VERSION : 1.2
// ellipse_C calculates the circumference of an ellipe based on the two radians R1 and R2
   VAR_INPUT
      R1 : Real;
      R2 : Real;
   END_VAR
BEGIN


   #ELLIPSE_C := "PI" * (3.0 * (#R1+#R2) - SQRT((3.0 * #R1 + #R2) * (3.0 * #R2 + #R1)));


   (* revision histroy
   hm  16. oct 2007    rev 1.0
       original version

   hm  18. oct. 2008   rev 1.1
       using math constants

   hm  10. mar. 2009   rev 1.2
       changed syntax of real constants to 0.0

   *)
END_FUNCTION

FUNCTION "SPHERE_V" : Real   // FC160, SCL
TITLE = SPHERE_V
{ S7_Optimized_Access := 'FALSE' }
AUTHOR : hugo
FAMILY : GEOMETRY
NAME : SPHERE_V
VERSION : 1.2
// sphere_V calculates the Volume of a Sphere
   VAR_INPUT
      rx : Real;
   END_VAR
BEGIN


     #SPHERE_V := 4.188790205 * #rx * #rx * #rx;

   (* revision histroy
   hm  16. oct 2007  rev 1.0
     original version

   hm  4. dec 2007   rev 1.1
     changed code for better performance

   hm  22. feb 2008    rev 1.2
     changed code for better performance
   *)
END_FUNCTION

FUNCTION "TRIANGLE_A" : Real   // FC161, SCL
TITLE = TRIANGLE_A
{ S7_Optimized_Access := 'FALSE' }
AUTHOR : hugo
FAMILY : GEOMETRY
NAME : TRIANG_A
VERSION : 1.2
// triangle_A calculates the Area of a triangle.
// if any input is 0 it will be neglected and the are will be calculated from eiter:
// two sides and an angle (s1 and S2 and the angle A1) or 3 sides.
// 
// uses: RAD [FC100]
//       MODR [FC97] 
//       FLOOR2 [FC82]
   VAR_INPUT
      S1 : Real;
      "A" : Real;
      S2 : Real;
      S3 : Real;
   END_VAR
BEGIN


   IF #"A" = 0.0 THEN
       #TRIANGLE_A := SQRT((#S1+#S2+#S3) * (#S1+#S2-#S3) * (#S2+#S3-#S1) * (#S3+#S1-#S2)) * 0.25;
   ELSE
       #TRIANGLE_A := #S1 * #S2 * SIN("RAD"(#"A")) * 0.5;
   END_IF;


   (* revision histroy
   hm  16. oct 2007    rev 1.0
       original version

   hm  22. feb 2008    rev 1.1
       improved performance

   hm  10. mar. 2009   rev 1.2
       changed syntax of real constants to 0.0

   *)
END_FUNCTION

FUNCTION "CIRCLE_SEG" : Real   // FC428, SCL
TITLE = CIRCLE_SEG
{ S7_Optimized_Access := 'FALSE' }
AUTHOR : hugo
FAMILY : GEOMETRY
NAME : CIRCLSEG
VERSION : 1.0
// CIRCLE_SEG calculates the Area of a circle segement enclosed between a sectant line and the circumference.
   VAR_INPUT
      RX : Real;
      HX : Real;
   END_VAR
BEGIN


   IF #RX > 0.0 THEN
     #CIRCLE_SEG := 2.0 * ACOS(1.0 - LIMIT(MN:=0.0,IN:=#HX / #RX,MX:=2.0));
     #CIRCLE_SEG := (#CIRCLE_SEG - SIN(#CIRCLE_SEG)) *#RX * #RX / 2.0;
   END_IF;


   (* revision histroy
   hm  10. mar 2010  rev 1.0
     original version

   *)
END_FUNCTION

// ===== PLC "Mathematical functions"  Unspecific CPU S7 300 =====

VAR_GLOBAL CONSTANT   // PLC tag table "STEP7 classic symbols"
   "debug" : Bool := FALSE;
   "N" : Int := 0;
   "offset" : Int := 0;
   "offset_1" : DWord := 0;
END_VAR

TYPE "XY_LINEAR_INT"
VERSION : 0.0
   STRUCT
      XY : Array[1..20, 0..1] of Real;
   END_STRUCT;
END_TYPE

TYPE "XY_POLYNOM_INT"
VERSION : 0.0
   STRUCT
      XY : Array[1..5, 0..1] of Real;
   END_STRUCT;
END_TYPE

TYPE "C_F_POLY"
VERSION : 0.0
   STRUCT
      C : Array[0..7] of Real;
   END_STRUCT;
END_TYPE

DATA_BLOCK "IDB_STIME"   // DB64
{ S7_Optimized_Access := 'FALSE' }
AUTHOR : dalbi
FAMILY : MEASURE
VERSION : 0.0
// stored: InstanceOfName STIME
"STIME"
BEGIN
END_DATA_BLOCK

FUNCTION_BLOCK "FT_AVG"   // FB23, SCL
TITLE = FT_AVG
{ S7_Optimized_Access := 'FALSE' }
AUTHOR : hugo
FAMILY : FUNCT
NAME : FT_AVG
VERSION : 1.5
// this function calculates the average over n samples from a sequential input
// the input values are shifted into an N deep buffer and the avg of this buffer is diplayed at anytime on the output.
// a rst will load the buffer with the current in value..
//  
// uses: DELAY [FB107]
//       INC1 [FC53]
   VAR_INPUT
      IN : Real;
      "E" : Bool := TRUE;
      N : Int := 32;
      RST : Bool;
   END_VAR
   VAR_OUTPUT
      AVG : Real;
   END_VAR
   VAR
      buff : "DELAY";
      i : Int;
      init : Bool;
   END_VAR
BEGIN


   (* limit n to a max of 32 because delay can do max 32 cycles *)
   #buff.N := LIMIT(MN:=0,IN:=#N,MX:=32);

   IF NOT #init OR #RST THEN
       FOR #i := 1 TO #N DO
           #buff(IN := #IN);
       END_FOR;
       #AVG := #IN;
       #init := TRUE;
   ELSIF #"E" THEN
       #buff(IN := #IN);
       #AVG := #AVG + (#IN - #buff.OUT) / INT_TO_REAL(#N);
   END_IF;


   (* revision history

   hm  7. jan. 2007    rev 1.1
       chaged rst logic to load the buffer with the actual input value instead of 0.
       added en input to allow better control of signal flow
       added init to load the buffer with in at startup to avoid rampup at beginning.
       deleted unused variable cnt.

   hm  14. jun. 2008   rev 1.2
       set default for input en = TRUE and N = 32

   hm  10. oct. 2008   rev 1.3
       improved performance

   hm  18. oct. 2008   rev 1.4
       changed input en to e for compatibility reasons

   hm  10. mar. 2009   rev 1.5
       added type conversion for compatibility reasons

   *)
END_FUNCTION_BLOCK

FUNCTION_BLOCK "FT_MIN_MAX"   // FB24, SCL
TITLE = FT_MIN_MAX
{ S7_Optimized_Access := 'FALSE' }
AUTHOR : hugo
FAMILY : FUNCT
NAME : MIN_MAX
VERSION : 1.0
// this function block stores the min and max value of an input signal.
// when rst is true the mn and mx outputs are set to the in value.
// when a rst is never active the function autoresets to the in value at startup.
// since the input might not be present at first cycle the mn and mx are set during second cycle.
   VAR_INPUT
      in : Real;
      rst : Bool;
   END_VAR
   VAR_OUTPUT
      mx : Real;
      mn : Real;
   END_VAR
   VAR
      init : Bool;
   END_VAR
BEGIN


     IF #rst OR NOT #init THEN
       #mn := #in;
       #mx := #in;
       #init := 1;
     ELSIF #in < #mn THEN
       #mn := #in;
     ELSIF #in > #mx THEN 
       #mx := #in;
     END_IF;
END_FUNCTION_BLOCK

FUNCTION_BLOCK "FT_RMP"   // FB25, SCL
TITLE = FT_RMP
{ S7_Optimized_Access := 'FALSE' }
AUTHOR : oscat
FAMILY : FUNCT
NAME : RMP
VERSION : 1.4
// this ramp function follows an input signal with a linear ramp up or down, the up or down speed can be set with KF and KR.
// a K factor of 1 means 1 unit per second on the output. K factors can only be positive and not negative.
// a busy output signals the ramp is running or busy false means the in value is present on the output.
// a rmp input false means the output follows the input dierctly while a rmp = true means the output follows the input with a ramp.
// a updn output signal the directon of the ramp (up or down).
// 
// uses: T_PLC_MS [FC64]
//       STIME [FB64],IDB_STIME [DB64]
   VAR_INPUT
      Rmp : Bool := TRUE;
      in : Real;
      KR : Real;
      KF : Real;
   END_VAR
   VAR_OUTPUT
      out : Real;
      busy : Bool;
      UD : Bool;
   END_VAR
   VAR
      tx : Time;
      last : Time;
      init : Bool;
   END_VAR
BEGIN


     (* read system time *)
     #tx := T_CONV(DWORD_TO_DINT("T_PLC_MS"())) - #last;

     IF NOT #init THEN
       #init := TRUE;
       #last := #tx;
       #tx := t#0s;
       #out := #in;
     END_IF;
     IF NOT #Rmp THEN
       #out := #in;
       #busy := FALSE;
     ELSIF #out > #in THEN
       (* ramp down *)
       #out := #out - DINT_TO_REAL(T_CONV(#tx)) * 0.001 * #KF;
       #out := MAX(IN1:=#in,IN2:=#out);
     ELSIF #out < #in THEN
       (* ramp up *)
       #out := #out + DINT_TO_REAL(T_CONV(#tx)) * 0.001 * #KR;
       #out := MIN(IN1:=#in,IN2:=#out);
     END_IF;

     (* set busy and dir flags *)
     IF #out < #in THEN
       #busy := TRUE;
       #UD := 1;
     ELSIF #out > #in THEN
       #busy := TRUE;
       #UD := 0;
     ELSE
       #busy := FALSE;
     END_IF;
     #last := #last + #tx;


   (* revision history:

   hm 8.10.2006      rev 1.1
     added ud output

   hm 12. feb 2007   rev 1.2
     added init variable and corrected a possible startup problem

   hm  17. sep 2007  rev 1.3
     replaced time() with t_plc_ms() for compatibility reasons

   hm  25. jan 2008  rev 1.4
     performance improvements
     allow KR and KF to be 0
   *)
END_FUNCTION_BLOCK

FUNCTION_BLOCK "STIME"   // FB64, SCL
TITLE = STIME
{ S7_Optimized_Access := 'FALSE' }
AUTHOR : dalbi
FAMILY : MEASURE
NAME : STIME
VERSION : 1.4
// this function block makes sure that the timer of a siemens sps counts from 0 - 2^32-1.
   VAR_OUTPUT
      tx : DWord;
      at_tx AT tx : Array[0..31] of Bool;
   END_VAR
   VAR
      last_time : DWord;
      bit31 : Bool;
      init : Bool := TRUE;
   END_VAR
   VAR_TEMP
      TOP_SI : Struct
         EV_CLASS : Byte;
         EV_NUM : Byte;
         PRIORITY : Byte;
         NUM : Byte;
         TYP2_3 : Byte;
         TYP1 : Byte;
         ZI1 : Word;
         ZI2_3 : DWord;
      END_STRUCT;
      START_UP_SI : Struct
         EV_CLASS : Byte;
         EV_NUM : Byte;
         PRIORITY : Byte;
         NUM : Byte;
         TYP2_3 : Byte;
         TYP1 : Byte;
         ZI1 : Word;
         ZI2_3 : DWord;
      END_STRUCT;
      ERR : Int;
   END_VAR
BEGIN


   (* this FB is only necessary for siemens sps
   the siemens sps timer counts from 0 to 2^31-1 and starts at 0 sfter overrun.
   this means that the bit 31 (the highest bit ) will never be used and therefore
   a problem arises when t2 - t1 is checked.
   t2 - t1 is always valid also in an timer overrun situation where the time t1 is very high and t2 is very low.
   the result of the subtraction t2 - t1 however is still valid.
   this calculation does not work for soiemens because the highest bit is not used.

   this module stores the highest bit, changes the highest bit at every overrun occurence and stuffs ther highest bit in the output.
   the output is then used by t_plc_us and t_plc_ms.

   the correction needs and fb and not a function because the value of the highest bit has to be stored.

   do never use this function block in a codesys environment. the timer in codesys is correct and runs from 0 to 2^32-1
   *)

   (* read actual startup info *)
   (* OB1_SCAN_1  BYTE  -  B#16#01: Abschluss des Neustarts (Warmstarts)
                        -  B#16#02: Abschluss des Wiederanlaufs
                        -  B#16#03: Abschluss des freien Zyklus
                        -  B#16#04: Abschluss des Kaltstarts
                        -  B#16#05: Erster OB 1-Zyklus der neuen Master-CPU nach 
                                    Master-Reserve-Umschaltung und STOP des 
                                    bisherigen Masters *)

   #ERR := RD_SINFO (TOP_SI => #TOP_SI, START_UP_SI => #START_UP_SI);

   (* reset last_time on system startup *)
   IF #TOP_SI.EV_NUM = 1 OR #TOP_SI.EV_NUM = 2 OR #TOP_SI.EV_NUM = 4 OR NOT #init THEN 
       #last_time := 0;
       #bit31 := false;
       #init := true;
   END_IF;

   (* read the system timer *)
   #tx := DINT_TO_DWORD(T_CONV(TIME_TCK()));

   (* check for overrun *)
   IF DWORD_TO_DINT(#tx) < DWORD_TO_DINT(#last_time) THEN
       (* an overrun has occured, change the value of the highest bit *)
       #bit31 := NOT #bit31;
   END_IF;

   (* stuff the highest bit into the timer value *)
   #at_tx[7] := #bit31;

   (* remember the last system time for the next overrun check *)
   #last_time := #tx;


   (* revision history
   DA  14.9.2007 rev 1.0
     original version

   DA  24.2.2008 rev 1.1
     added self reset on system startup

   DA   2.5.2008 rev 1.2
     corect a problem running under OB35

   DA  12.3.2009 rev 1.3
     corect a problem run on different CPUs

   DA  22.12.2009 rev 1.4
     corect a problem on startup
   *)
END_FUNCTION_BLOCK

FUNCTION_BLOCK "DELAY"   // FB107, SCL
TITLE = DELAY
{ S7_Optimized_Access := 'FALSE' }
AUTHOR : hugo
FAMILY : SIGPRO
NAME : DELAY
VERSION : 1.5
// this function block delays input values by each programm cycle
// after N+1 cycles the in value has shifted to the out.
// N can be any alue from 0 .. 32
// if n = 0 the input will be present on the output without a delay.
// f N > 32 then the output will be delayed by 32 cycles.
// any high on rst will load the buffer with in.
// 
// uses: INC1 [FC53]
   VAR_INPUT
      IN : Real;
      N : Int;
      RST : Bool;
   END_VAR
   VAR_OUTPUT
      OUT : Real;
   END_VAR
   VAR
      buf : Array[0..31] of Real;
      i : Int;
      init : Bool;
      stop : Int;
   END_VAR
BEGIN


   #stop := LIMIT(MN:=0,IN:=#N,MX:=32) - 1;
   IF #RST OR NOT #init THEN
       #init := TRUE;
       FOR #i := 0 TO #stop DO #buf[#i] := #IN; END_FOR;
       #OUT := #IN;
       #i := 0;         // Muss so sein!
   ELSIF #stop < 0 THEN
       #OUT := #IN;
   ELSE
       #OUT := #buf[#i];
       #buf[#i] := #IN;
       #i := "INC1"(X:=#i, N:=#N);
   END_IF;


   (* revision history
   hm 1.10.2006        rev 1.1
       corrected error in buffer management

   hm 19.1.2007        rev 1.2
       changed reset to load the value of in instead of 0

   hm  27. oct. 2008   rev 1.3
       improved performance

   hm  23. feb.2009    rev 1.4
       corrected an index problem

   hm  23. mar. 2009   rev 1.5
       corrected non standard write to input N

   *)
END_FUNCTION_BLOCK

FUNCTION "INC1" : Int   // FC53, SCL
TITLE = INC1
{ S7_Optimized_Access := 'FALSE' }
AUTHOR : hugo
FAMILY : MATH
NAME : INC1
VERSION : 1.2
// This is a increment function which increments the variable X by 1 and if M is reached, it begins with 0 again.
// _inc1(3,X) will generate 0,1,2,3,0,1,.....
   VAR_INPUT
      X : Int;
      N : Int;
   END_VAR
BEGIN


   IF #X >= #N - 1 THEN
       #INC1 := 0;
   ELSE
       #INC1 := #X + 1;
   END_IF;


   (* this elegant version is 50% slower
   INC1 := X := (x + 1) MOD N;
   *)



   (* revision history
   hm  13. oct. 2008   rev 1.0
       original version

   hm  22. oct. 2008   rev 1.1
       added statement to return value for compatibility reasons

   hm  23. feb. 2009   rev 1.2
       when inc1 is called with X >= N inc will continue with 0
   *)
END_FUNCTION

FUNCTION "T_PLC_MS" : DWord   // FC64, SCL
TITLE = T_PLC_MS
{ S7_Optimized_Access := 'FALSE' }
AUTHOR : hugo
FAMILY : MEASURE
NAME : T_PLC_MS
VERSION : 1.2
// T_PLC_MS reads the internal PLC timer and return the time, it has the advantage to be able to set a debug mode 
// and speed up the counter to test the plc timer overrun which occurs every 50 days respectively 25 days at siemens S7
// this routine also allows to correct the behavior of s7 where the internal plc counter will not count all 32 bits.
// 
// uses: STIME [FB64],IDB_STIME [DB64]
BEGIN


   "IDB_STIME"(); 
   #T_PLC_MS := "IDB_STIME".tx; 
   (* hier muss die korrektur für step7 stattfinden
   plctime muss den vollen wertebereich von time ausnutzen:
   wenn bei step7 time -24tage bis plus 24 tage ist dann muss der timer auch beim überlauf auf -24tage springen 
   und auf keinen fall auf 0 !!!!
   für siemens muss ein weiterer fb im main eingebunden werden der sicherstellt das alle 32 bits durchgezählt werden.
   es kann nur ein fb sein den er muss sich das oberste (32te) bit merken.
   oder etwa spring s7 bei überlauf auf -24 tage????? dann wäre keine korrektur nötig.
   *)
   IF "debug" THEN
       #T_PLC_MS := DINT_TO_DWORD((DWORD_TO_DINT(SHL(IN:=#T_PLC_MS,N:="N") OR SHL(IN:=DWORD#1,N:="N"))-1) + DWORD_TO_DINT("offset_1"));
   END_IF;


   (* revision history
   hm  14.9.2007   rev 1.0
       original version

   hm  12. nov 2007    rev 1.1
       added temporaray variable tx because some compilers could not handle time() as an argument

   hm  16. nov. 2008   rev 1.2
       initialized constants with 0 for compatibility reasons
   *)
END_FUNCTION

FUNCTION "F_LIN" : Real   // FC148, SCL
TITLE = F_LIN
{ S7_Optimized_Access := 'FALSE' }
AUTHOR : hugo
FAMILY : FUNCT
NAME : LIN
VERSION : 1.0
// this function calculates the linear equation f_lin = a*x + b
   VAR_INPUT
      X : Real;
      "A" : Real;
      "B" : Real;
   END_VAR
BEGIN


     #F_LIN := #"A" * #X + #"B";
END_FUNCTION

FUNCTION "F_LIN2" : Real   // FC149, SCL
TITLE = F_LIN2
{ S7_Optimized_Access := 'FALSE' }
AUTHOR : hugo
FAMILY : FUNCT
NAME : LIN2
VERSION : 1.1
// this function calculates the linear equation f_lin = a*x + b given by two points x1/y1 and x2/y2.
   VAR_INPUT
      X : Real;
      X1 : Real;
      Y1 : Real;
      X2 : Real;
      Y2 : Real;
   END_VAR
BEGIN


   #F_LIN2 := (#Y2 - #Y1) / (#X2 - #X1) * (#X - #X1) + #Y1;


   (* revision history
   hm  1. jan. 2007    rev 1.0
       original release

   hm  17. dec. 2008   rev 1.1
       optimized formula

   *)
END_FUNCTION

FUNCTION "F_POLY" : Real   // FC150, SCL
TITLE = F_POLY
{ S7_Optimized_Access := 'FALSE' }
AUTHOR : hugo
FAMILY : FUNCT
NAME : F_POLY
VERSION : 1.1
// this function calculates the polynom C[0] + C[1]*X^1 + C[2]*X^2 * C[3]*X^3 + C[4]*X^4 + C[5]*X^5 + C[6]*X^6 + C[7]*X^7
// 
// uses: C_F_POLY [UDT18]
   VAR_INPUT
      X : Real;
      C : "C_F_POLY";
   END_VAR
   VAR_TEMP
      x2 : Real;
      X4 : Real;
      X6 : Real;
   END_VAR
BEGIN


   #F_POLY := ((((((( #C.C[7] * #X + #C.C[6] ) * #X + #C.C[5] ) * #X + #C.C[4] ) * #X + #C.C[3] ) * #X + #C.C[2] ) * #X + #C.C[1] ) * #X + #C.C[0] ) ;


   (* revision history
   hm    20. may. 2008   rev 1.0
     original version

   hm  18. mar. 2011 rev 1.1
     improved performance
   *)
END_FUNCTION

FUNCTION "F_POWER" : Real   // FC151, SCL
TITLE = F_POWER
{ S7_Optimized_Access := 'FALSE' }
AUTHOR : hugo
FAMILY : FUNCT
NAME : POWER
VERSION : 1.0
// this function calculates the power equation f_power = a*x^n
   VAR_INPUT
      "a" : Real;
      x : Real;
      n : Real;
   END_VAR
BEGIN


     #F_POWER := #"a" * (#x**#n);
END_FUNCTION

FUNCTION "F_QUAD" : Real   // FC152, SCL
TITLE = F_QUAD
{ S7_Optimized_Access := 'FALSE' }
AUTHOR : hugo
FAMILY : FUNCT
NAME : QUAD
VERSION : 1.1
// this function calculates the quadratic equation f_lin = a*x + b
   VAR_INPUT
      X : Real;
      "A" : Real;
      "B" : Real;
      C : Real;
   END_VAR
BEGIN


   #F_QUAD :=  (#"A" * #X + #"B") * #X + #C;


   (* revision history

   hm  1. sep. 2006  rev 1.0
     original version

   hm  18. mar. 2001 rev 1.1
     improved performance
   *)
END_FUNCTION

FUNCTION "LINEAR_INT" : Real   // FC153, SCL
TITLE = LINEAR_INT
{ S7_Optimized_Access := 'FALSE' }
AUTHOR : oscat
FAMILY : FUNCT
NAME : LIN_INT
VERSION : 1.1
// LINEAR_INT calculates an output based on a linear interpolation of up to 20 coordinates given in an array
// the indut coordinates have to start at the lowest array position and must be sorted ba ascending X values.
// 
// uses: XY_LINEAR_INT [UDT16]
   VAR_INPUT
      X : Real;
      XY : "XY_LINEAR_INT";
      Pts : Int;
   END_VAR
   VAR_TEMP
      temp_Pts : Int;
      i : Int;
   END_VAR
BEGIN


     #temp_Pts := #Pts;

   (* make sure n is bound within the array size *)
     #temp_Pts := MIN(IN1:=#temp_Pts,IN2:=20);

   (* calculate the linear segement interpolation *)
     #i := 2;
   (* search for segment and calculate output
     below and above the defined segments we interpolate the last segment *)
     WHILE (#i < #temp_Pts) AND (#XY.XY[#i,0] < #X) DO
       #i := #i + 1;
     END_WHILE;

   (* calculate the output value on the corresponding segment coordinates *)
     #LINEAR_INT := ((#XY.XY[#i,1] - #XY.XY[#i-1,1]) * #X - #XY.XY[#i,1] * #XY.XY[#i-1,0] + #XY.XY[#i-1,1]*#XY.XY[#i,0]) / (#XY.XY[#i,0] - #XY.XY[#i-1,0]);

   (* revision history
   hm  7. oct 2007   rev 1.0
     original version

   hm  27 dec 2007   rev 1.1
     changed code for better performance
   *)
END_FUNCTION

FUNCTION "POLYNOM_INT" : Real   // FC154, SCL
TITLE = POLYNOM_INT
{ S7_Optimized_Access := 'FALSE' }
AUTHOR : oscat
FAMILY : FUNCT
NAME : POLY_INT
VERSION : 1.3
// POLYNOM_INT calculates an output based on a Polynom interpolation of up to 5 coordinates given in an array
// the indut coordinates have to start at the lowest array position and must be sorted ba ascending X values.
// 
// uses: XY_POLYNOM_INT [UDT17]
   VAR_INPUT
      X : Real;
      XY : "XY_POLYNOM_INT";
      Pts : Int;
   END_VAR
   VAR_TEMP
      I : Int;
      J : Int;
      stop : Int;
      tPts : Int;
      tXY : "XY_POLYNOM_INT";
   END_VAR
BEGIN


   #tXY := #XY;
   #tPts := #Pts;

   (* make sure n is bound within the array size *)
   #tPts := MIN(IN1:=#tPts,IN2:=5);

   (* this part is only to calculate the polynom parameters, which are then stores in the Y array
     the array values, it is not needed during runtime, unless the parameters will change during runtime
     the remaining code without this setup code can be used within a function to calculate specific functions
     the content of the arrays is then used as constant values within the function *)

   FOR #I := 1 TO #tPts DO
       #stop := #I + 1;
       FOR #J := #tPts TO #stop BY -1 DO
           #tXY.XY[#J,1] := (#tXY.XY[#J,1] - #tXY.XY[#J-1,1]) / (#tXY.XY[#J,0] - #tXY.XY[#J-#I,0]);
       END_FOR;
   END_FOR;


   (* this part is the actual calculation *)
   #POLYNOM_INT := 0.0;
   FOR #I := #tPts TO 1 BY -1 DO
          #POLYNOM_INT := #POLYNOM_INT * (#X - #tXY.XY[#I,0]) + #tXY.XY[#I,1];
   END_FOR;


   (* revision history
   hm  8. okt 2007 rev 1.0
       original version

   hm  17. dec 2007    rev 1.1
       init makes no sense for a function

   hm  22. feb 2008    rev 1.2
       improved performance

   hm  10. mar. 2009   rev 1.3
       changed syntax of real constants to 0.0

   *)
END_FUNCTION

FUNCTION "FRMP_B" : Byte   // FC424, SCL
TITLE = FRMP_B
{ S7_Optimized_Access := 'FALSE' }
AUTHOR : hugo
FAMILY : FUNCT
NAME : FRMP_B
VERSION : 1.0
// this function calculates a ramp and limits the output to 0 .. 255 without overflow problems
   VAR_INPUT
      START : Byte;
      DIR : Bool;
      TD : Time;
      TR : Time;
   END_VAR
   VAR_TEMP
      tTD : Time;
   END_VAR
BEGIN


   #tTD := #TD;  // only Step7

   IF #TD < #TR THEN
     #FRMP_B := DINT_TO_BYTE(MIN(IN1:=DWORD_TO_DINT(SHL(IN:=DINT_TO_DWORD(T_CONV(#tTD)), N:=8)) / T_CONV(#TR) 
                                ,IN2:=SEL(G:=#DIR, IN0:=BYTE_TO_DINT(#START), IN1:=BYTE_TO_DINT(BYTE#255) - BYTE_TO_DINT(#START))));
     IF #DIR THEN
       #FRMP_B := INT_TO_BYTE(BYTE_TO_INT(#START) + BYTE_TO_INT(#FRMP_B));
     ELSE
       #FRMP_B := INT_TO_BYTE(BYTE_TO_INT(#START) - BYTE_TO_INT(#FRMP_B));
     END_IF;
   ELSE
     #FRMP_B := INT_TO_BYTE(IN:= DINT_TO_INT(IN:= SEL(G:=#DIR, IN0:=0, IN1:=255)));
   END_IF;


   (* revision history

   17. feb. 2011 rev 1.0
     new module

   *)
END_FUNCTION

// ===== PLC "Other"  Unspecific CPU S7 300 =====

VAR_GLOBAL CONSTANT   // PLC tag table "STEP7 classic symbols"
   "debug" : Bool := FALSE;
   "N" : Int := 0;
   "offset" : Int := 0;
   "offset_1" : DWord := 0;
END_VAR

TYPE "ESR_DATA"
VERSION : 0.0
   STRUCT
      TYP : Byte;
      ADRESS : String[10];
      DS : Date_And_Time;
      TS : Time;
      DATA : Array[0..7] of Byte;
   END_STRUCT;
END_TYPE

DATA_BLOCK "IDB_STIME"   // DB64
{ S7_Optimized_Access := 'FALSE' }
AUTHOR : dalbi
FAMILY : MEASURE
VERSION : 0.0
// stored: InstanceOfName STIME
"STIME"
BEGIN
END_DATA_BLOCK

FUNCTION_BLOCK "ESR_COLLECT"   // FB1, SCL
TITLE = ESR_COLLECT
{ S7_Optimized_Access := 'FALSE' }
AUTHOR : hugo
FAMILY : OTHER
NAME : ESR_COLL
VERSION : 1.4
// ESR_collect collects esr data from up to 8 esr_mon modules and stroes them in an output array.
//  the output pos will display the position of the last element in the array. if the array is empty, pos = -1
//  when to buffer is read by followon modules. pos has to be reset to -1
//  if the array will be full, the buffer will be refilled starting at position 0.
// 
// uses: ESR_DATA [UDT8]
//       INC1 [FC53]
   VAR_INPUT
      ESR_0 : Array[0..3] of "ESR_DATA";
      ESR_1 : Array[0..3] of "ESR_DATA";
      ESR_2 : Array[0..3] of "ESR_DATA";
      ESR_3 : Array[0..3] of "ESR_DATA";
      ESR_4 : Array[0..3] of "ESR_DATA";
      ESR_5 : Array[0..3] of "ESR_DATA";
      ESR_6 : Array[0..3] of "ESR_DATA";
      ESR_7 : Array[0..3] of "ESR_DATA";
      RST : Bool;
   END_VAR
   VAR_OUTPUT
      ESR_OUT : Array[0..31] of "ESR_DATA";
   END_VAR
   VAR_IN_OUT
      pos : Int;
   END_VAR
   VAR
      max_in : Int := 3;
      max_out : Int := 32;
      cnt : Int := -1;
   END_VAR
BEGIN


   IF #RST OR #cnt < 0 THEN
     #pos := -1;
   ELSE
     FOR #cnt := 0 TO #max_in DO
       IF BYTE_TO_INT(#ESR_0[#cnt].TYP) > 0 THEN #pos := "INC1"(X:=#pos, N:=#max_out); #ESR_OUT[#pos] := #ESR_0[#cnt]; END_IF;
       IF BYTE_TO_INT(#ESR_1[#cnt].TYP) > 0 THEN #pos := "INC1"(X:=#pos, N:=#max_out); #ESR_OUT[#pos] := #ESR_1[#cnt]; END_IF;
       IF BYTE_TO_INT(#ESR_2[#cnt].TYP) > 0 THEN #pos := "INC1"(X:=#pos, N:=#max_out); #ESR_OUT[#pos] := #ESR_2[#cnt]; END_IF;
       IF BYTE_TO_INT(#ESR_3[#cnt].TYP) > 0 THEN #pos := "INC1"(X:=#pos, N:=#max_out); #ESR_OUT[#pos] := #ESR_3[#cnt]; END_IF;
       IF BYTE_TO_INT(#ESR_4[#cnt].TYP) > 0 THEN #pos := "INC1"(X:=#pos, N:=#max_out); #ESR_OUT[#pos] := #ESR_4[#cnt]; END_IF;
       IF BYTE_TO_INT(#ESR_5[#cnt].TYP) > 0 THEN #pos := "INC1"(X:=#pos, N:=#max_out); #ESR_OUT[#pos] := #ESR_5[#cnt]; END_IF;
       IF BYTE_TO_INT(#ESR_6[#cnt].TYP) > 0 THEN #pos := "INC1"(X:=#pos, N:=#max_out); #ESR_OUT[#pos] := #ESR_6[#cnt]; END_IF;
       IF BYTE_TO_INT(#ESR_7[#cnt].TYP) > 0 THEN #pos := "INC1"(X:=#pos, N:=#max_out); #ESR_OUT[#pos] := #ESR_7[#cnt]; END_IF;
     END_FOR;
   END_IF;


   (* revision history
   hm  26.jan 2007 rev 1.0
     original version

   hm  8. dec 2007 rev 1.1
     added reset input

   ks  27. oct. 2008 rev 1.2
     optimized code for performance

   ks  12. nov. 2009 rev 1.3
     output pos was not pointing to last value 

   hm  1. dec. 2009 rev 1.4
     changed pos to be I/O
     reduced output array size to 32 elements
   *)
END_FUNCTION_BLOCK

FUNCTION_BLOCK "ESR_MON_B8"   // FB2, SCL
TITLE = ESR_MON_B8
{ S7_Optimized_Access := 'FALSE' }
AUTHOR : hugo
FAMILY : OTHER
NAME : ESRMONB8
VERSION : 1.3
// ESR_mon_B8 monitores up to 8 binary inputs and reports changes with time stamd and adress label.
// the module checks 8 inputs for a change and reports all changes with time and adress stamp to the output.
// 4 events maximum can be collected at once within the same cycle
// 
// uses: ESR_DATA [UDT8]
//       T_PLC_MS [FC64]
//       STIME [FB64],IDB_STIME [DB64]
   VAR_INPUT
      s0 : Bool;
      s1 : Bool;
      s2 : Bool;
      s3 : Bool;
      s4 : Bool;
      s5 : Bool;
      s6 : Bool;
      s7 : Bool;
      DT_in : Date_And_Time;
      a0 : String[10];
      a1 : String[10];
      a2 : String[10];
      a3 : String[10];
      a4 : String[10];
      a5 : String[10];
      a6 : String[10];
      a7 : String[10];
   END_VAR
   VAR_OUTPUT
      ESR_Flag : Bool;
   END_VAR
   VAR_IN_OUT
      ESR_Out : Array[0..3] of "ESR_DATA";
   END_VAR
   VAR
      x0 : Bool;
      x1 : Bool;
      x2 : Bool;
      x3 : Bool;
      x4 : Bool;
      x5 : Bool;
      x6 : Bool;
      x7 : Bool;
      tx : Time;
      cnt : Int;
   END_VAR
BEGIN


   (* read system timer *)
   #tx := T_CONV(DWORD_TO_DINT("T_PLC_MS"()));

   #ESR_Flag := FALSE;
   #ESR_Out[3].TYP := 0;
   #ESR_Out[2].TYP := 0;
   #ESR_Out[1].TYP := 0;
   #ESR_Out[0].TYP := 0;
   #cnt := 0;

   (* check if inputs have chaged and fill buffer *)
   IF #s0 <> #x0 THEN
       #ESR_Out[#cnt].TYP := INT_TO_BYTE(10 + BOOL_TO_INT(#s0));
       #ESR_Out[#cnt].ADRESS := #a0;
       #ESR_Out[#cnt].DS := #DT_in;
       #ESR_Out[#cnt].TS := #tx;
       #x0 := #s0;
       #cnt := #cnt + 1;
       #ESR_Flag := TRUE;
   END_IF;
   IF #s1 <> #x1 THEN
       #ESR_Out[#cnt].TYP := INT_TO_BYTE(10 + BOOL_TO_INT(#s1));
       #ESR_Out[#cnt].ADRESS BLKMOV #a1;
       #ESR_Out[#cnt].DS := #DT_in;
       #ESR_Out[#cnt].TS := #tx;
       #x1 := #s1;
       #cnt := #cnt + 1;
       #ESR_Flag := TRUE;
   END_IF;
   IF #s2 <> #x2 THEN
       #ESR_Out[#cnt].TYP := INT_TO_BYTE(10 + BOOL_TO_INT(#s2));
       #ESR_Out[#cnt].ADRESS BLKMOV #a2;
       #ESR_Out[#cnt].DS := #DT_in;
       #ESR_Out[#cnt].TS := #tx;
       #x2 := #s2;
       #cnt := #cnt + 1;
       #ESR_Flag := TRUE;
   END_IF;
   IF #s3 <> #x3 THEN
       #ESR_Out[#cnt].TYP := INT_TO_BYTE(10 + BOOL_TO_INT(#s3));
       #ESR_Out[#cnt].ADRESS BLKMOV #a3;
       #ESR_Out[#cnt].DS := #DT_in;
       #ESR_Out[#cnt].TS := #tx;
       #x3 := #s3;
       #cnt := #cnt + 1;
       #ESR_Flag := TRUE;
   END_IF;
   IF #s4 <> #x4 AND #cnt < 4 THEN
       #ESR_Out[#cnt].TYP := INT_TO_BYTE(10 + BOOL_TO_INT(#s4));
       #ESR_Out[#cnt].ADRESS BLKMOV #a4;
       #ESR_Out[#cnt].DS := #DT_in;
       #ESR_Out[#cnt].TS := #tx;
       #x4 := #s4;
       #cnt := #cnt + 1;
       #ESR_Flag := TRUE;
   END_IF;
   IF #s5 <> #x5  AND #cnt < 4 THEN
       #ESR_Out[#cnt].TYP := INT_TO_BYTE(10 + BOOL_TO_INT(#s5));
       #ESR_Out[#cnt].ADRESS BLKMOV #a5;
       #ESR_Out[#cnt].DS := #DT_in;
       #ESR_Out[#cnt].TS := #tx;
       #x5 := #s5;
       #cnt := #cnt + 1;
       #ESR_Flag := TRUE;
   END_IF;
   IF #s6 <> #x6  AND #cnt < 4 THEN
       #ESR_Out[#cnt].TYP := INT_TO_BYTE(10 + BOOL_TO_INT(#s6));
       #ESR_Out[#cnt].ADRESS BLKMOV #a6;
       #ESR_Out[#cnt].DS := #DT_in;
       #ESR_Out[#cnt].TS := #tx;
       #x6 := #s6;
       #cnt := #cnt + 1;
       #ESR_Flag := TRUE;
   END_IF;
   IF #s7 <> #x7  AND #cnt < 4 THEN
       #ESR_Out[#cnt].TYP := INT_TO_BYTE(10 + BOOL_TO_INT(#s7));
       #ESR_Out[#cnt].ADRESS BLKMOV #a7;
       #ESR_Out[#cnt].DS := #DT_in;
       #ESR_Out[#cnt].TS := #tx;
       #x7 := #s7;
       #cnt := #cnt + 1;
       #ESR_Flag := TRUE;
   END_IF;


   (* revision history
   hm  26. jan 2007  rev 1.0
     original version

   hm  17. sep 2007  rev 1.1
     replaced time() with T_PLC_MS() for compatibility reasons

   hm  22. oct. 2008 rev 1.2
     optimized code

   hm  1.dec. 2009 rev 1.3
     changed esr_out to be I/O

   *)
END_FUNCTION_BLOCK

FUNCTION_BLOCK "ESR_MON_R4"   // FB3, SCL
TITLE = ESR_MON_R4
{ S7_Optimized_Access := 'FALSE' }
AUTHOR : hugo
FAMILY : OTHER
NAME : ESRMONR4
VERSION : 1.4
// ESR_mon_R4 monitores up to 4 Real inputs and reports changes with time stamd and adress label.
// the module checks 4 inputs for a change of more than the specified sensitivity S and reports all changes with time and adress stamp to the output.
//  
// uses: ESR_DATA [UDT8]
//       T_PLC_MS [FC64]
//       STIME [FB64],IDB_STIME [DB64]
//       DIFFER [FC73]
   VAR_INPUT
      R0 : Real;
      p0 AT R0 : Array[0..3] of Byte;
      R1 : Real;
      p1 AT R1 : Array[0..3] of Byte;
      R2 : Real;
      p2 AT R2 : Array[0..3] of Byte;
      R3 : Real;
      p3 AT R3 : Array[0..3] of Byte;
      DT_in : Date_And_Time;
      a0 : String[10];
      a1 : String[10];
      a2 : String[10];
      a3 : String[10];
      s0 : Real;
      s1 : Real;
      s2 : Real;
      s3 : Real;
   END_VAR
   VAR_OUTPUT
      ESR_Flag : Bool;
   END_VAR
   VAR_IN_OUT
      ESR_Out : Array[0..3] of "ESR_DATA";
   END_VAR
   VAR
      x0 : Real;
      x1 : Real;
      x2 : Real;
      x3 : Real;
      tx : Time;
      cnt : Int;
   END_VAR
BEGIN


     (* read system timer *)
     #tx := T_CONV(DWORD_TO_DINT("T_PLC_MS"()));
     #ESR_Flag := FALSE;
     #ESR_Out[3].TYP := 0;
     #ESR_Out[2].TYP := 0;
     #ESR_Out[1].TYP := 0;
     #ESR_Out[0].TYP := 0;
     #cnt := 0;

     (* check if inputs have chaged and fill buffer *)
     IF "DIFFER"(in1:=#R0, in2:=#x0, X:=#s0) THEN
         #ESR_Out[#cnt].TYP := 20;
         #ESR_Out[#cnt].ADRESS BLKMOV #a0;
         #ESR_Out[#cnt].DS := #DT_in;
         #ESR_Out[#cnt].TS := #tx;
         #ESR_Out[#cnt].DATA[0] := #p0[0];
         #ESR_Out[#cnt].DATA[1] := #p0[1];
         #ESR_Out[#cnt].DATA[2] := #p0[2];
         #ESR_Out[#cnt].DATA[3] := #p0[3];
         #x0 := #R0;
         #cnt := #cnt + 1;
         #ESR_Flag := TRUE;
     END_IF;
     IF "DIFFER"(in1:=#R1, in2:=#x1, X:=#s1) THEN
         #ESR_Out[#cnt].TYP := 20;
         #ESR_Out[#cnt].ADRESS BLKMOV #a1;
         #ESR_Out[#cnt].DS := #DT_in;
         #ESR_Out[#cnt].TS := #tx;
         #ESR_Out[#cnt].DATA[0] := #p1[0];
         #ESR_Out[#cnt].DATA[1] := #p1[1];
         #ESR_Out[#cnt].DATA[2] := #p1[2];
         #ESR_Out[#cnt].DATA[3] := #p1[3];
         #x1 := #R1;
         #cnt := #cnt + 1;
         #ESR_Flag := TRUE;
     END_IF;
     IF "DIFFER"(in1:=#R2, in2:=#x2, X:=#s2) THEN
         #ESR_Out[#cnt].TYP := 20;
         #ESR_Out[#cnt].ADRESS BLKMOV #a2;
         #ESR_Out[#cnt].DS := #DT_in;
         #ESR_Out[#cnt].TS := #tx;
         #ESR_Out[#cnt].DATA[0] := #p2[0];
         #ESR_Out[#cnt].DATA[1] := #p2[1];
         #ESR_Out[#cnt].DATA[2] := #p2[2];
         #ESR_Out[#cnt].DATA[3] := #p2[3];
         #x2 := #R2;
         #cnt := #cnt + 1;
         #ESR_Flag := TRUE;
     END_IF;
     IF "DIFFER"(in1:=#R3, in2:=#x3, X:=#s3) THEN
         #ESR_Out[#cnt].TYP := 20;
         #ESR_Out[#cnt].ADRESS BLKMOV #a3;
         #ESR_Out[#cnt].DS := #DT_in;
         #ESR_Out[#cnt].TS := #tx;
         #ESR_Out[#cnt].DATA[0] := #p3[0];
         #ESR_Out[#cnt].DATA[1] := #p3[1];
         #ESR_Out[#cnt].DATA[2] := #p3[2];
         #ESR_Out[#cnt].DATA[3] := #p3[3];
         #x3 := #R3;
         #cnt := #cnt + 1;
         #ESR_Flag := TRUE;
     END_IF;


   (* revision history
   hm  26. jan 2007  rev 1.0
     original version

   hm  17. sep. 2007   rev 1.1
     replaced time() with T_PLC_MS() for compatibility reasons

   hm  8. dec. 2007    rev 1.2
     corrected an error while esr typ would not be set

   hm  16. mar. 2008   rev 1.3
     deleted wrong conversion real_to_dword

   hm  1. dec 2009   rev 1.4
     changed esr_out to be I/O

   *)
END_FUNCTION_BLOCK

FUNCTION_BLOCK "ESR_MON_X8"   // FB4, SCL
TITLE = ESR_MON_X8
{ S7_Optimized_Access := 'FALSE' }
AUTHOR : hugo
FAMILY : OTHER
NAME : ESRMONX8
VERSION : 1.2
// ESR_MON_X8 is a status and error collector.
// the module checks 8 status inputs for a change and reports up to 4 input changes with time and adress stamp to the output.
// the mode can be 
// 1 for error only
// 2 for error and status
// 3 for error, status and debug
// the adress label of the 8 inputs can be configured individually.
// 
// uses: ESR_DATA [UDT8]
//       T_PLC_MS [FC64]
//       STIME [FB64],IDB_STIME [DB64]
//       STATUS_TO_ESR [FC51]
   VAR_INPUT
      s0 : Byte;
      s1 : Byte;
      s2 : Byte;
      s3 : Byte;
      s4 : Byte;
      s5 : Byte;
      s6 : Byte;
      s7 : Byte;
      DT_in : Date_And_Time;
      Mode : Byte := B#16#3;
      a0 : String[10];
      a1 : String[10];
      a2 : String[10];
      a3 : String[10];
      a4 : String[10];
      a5 : String[10];
      a6 : String[10];
      a7 : String[10];
   END_VAR
   VAR_OUTPUT
      ESR_Flag : Bool;
   END_VAR
   VAR_IN_OUT
      ESR_Out : Array[0..3] of "ESR_DATA";
   END_VAR
   VAR
      x0 : Byte;
      x1 : Byte;
      x2 : Byte;
      x3 : Byte;
      x4 : Byte;
      x5 : Byte;
      x6 : Byte;
      x7 : Byte;
      tx : Time;
      cnt : Int;
   END_VAR
BEGIN


     (* read system timer *)
     #tx := T_CONV(DWORD_TO_DINT("T_PLC_MS"()));

     #ESR_Flag := FALSE;
     #ESR_Out[3].TYP := 0;
     #ESR_Out[2].TYP := 0;
     #ESR_Out[1].TYP := 0;
     #ESR_Out[0].TYP := 0;
     #cnt := 0;

     (* check if inputs have chaged and fill buffer *)
     IF #s0 <> #x0 AND ((BYTE_TO_INT(#s0) < 100) OR (BYTE_TO_INT(#s0) > 99 AND BYTE_TO_INT(#s0) < 200 AND BYTE_TO_INT(#Mode) >= 2) OR (BYTE_TO_INT(#s0) > 199 AND #Mode = 3)) THEN
         #ESR_Out[#cnt] := "STATUS_TO_ESR"(status:=#s0,adress:=#a0,DT_in:=#DT_in,TS:=#tx);
         #x0 := #s0;
         #cnt := #cnt + 1;
         #ESR_Flag := TRUE;
     END_IF;
     IF #s1 <> #x1 AND ((BYTE_TO_INT(#s1) < 100) OR (BYTE_TO_INT(#s1) > 99 AND BYTE_TO_INT(#s1) < 200 AND BYTE_TO_INT(#Mode) >= 2) OR (BYTE_TO_INT(#s1) > 199 AND #Mode = 3)) THEN
         #ESR_Out[#cnt] := "STATUS_TO_ESR"(status:=#s1,adress:=#a1,DT_in:=#DT_in,TS:=#tx);
         #x1 := #s1;
         #cnt := #cnt + 1;
         #ESR_Flag := TRUE;
     END_IF;
     IF #s2 <> #x2 AND ((BYTE_TO_INT(#s2) < 100) OR (BYTE_TO_INT(#s2) > 99 AND BYTE_TO_INT(#s2) < 200 AND BYTE_TO_INT(#Mode) >= 2) OR (BYTE_TO_INT(#s2) > 199 AND #Mode = 3)) THEN
         #ESR_Out[#cnt] := "STATUS_TO_ESR"(status:=#s2,adress:=#a2,DT_in:=#DT_in,TS:=#tx);
         #x2 := #s2;
         #cnt := #cnt + 1;
         #ESR_Flag := TRUE;
     END_IF;
     IF #s3 <> #x3 AND ((BYTE_TO_INT(#s3) < 100) OR (BYTE_TO_INT(#s3) > 99 AND BYTE_TO_INT(#s3) < 200 AND BYTE_TO_INT(#Mode) >= 2) OR (BYTE_TO_INT(#s3) > 199 AND #Mode = 3)) THEN
         #ESR_Out[#cnt] := "STATUS_TO_ESR"(status:=#s3,adress:=#a3,DT_in:=#DT_in,TS:=#tx);
         #x3 := #s3;
         #cnt := #cnt + 1;
         #ESR_Flag := TRUE;
     END_IF;
     IF #cnt < 4 AND #s4 <> #x4 AND ((BYTE_TO_INT(#s4) < 100) OR (BYTE_TO_INT(#s4) > 99 AND BYTE_TO_INT(#s4) < 200 AND BYTE_TO_INT(#Mode) >= 2) OR (BYTE_TO_INT(#s4) > 199 AND #Mode = 3)) THEN
         #ESR_Out[#cnt] := "STATUS_TO_ESR"(status:=#s4,adress:=#a4,DT_in:=#DT_in,TS:=#tx);
         #x4 := #s4;
         #cnt := #cnt + 1;
         #ESR_Flag := TRUE;
     END_IF;
     IF #cnt < 4 AND #s5 <> #x5 AND ((BYTE_TO_INT(#s5) < 100) OR (BYTE_TO_INT(#s5) > 99 AND BYTE_TO_INT(#s5) < 200 AND BYTE_TO_INT(#Mode) >= 2) OR (BYTE_TO_INT(#s5) > 199 AND #Mode = 3)) THEN
         #ESR_Out[#cnt] := "STATUS_TO_ESR"(status:=#s5,adress:=#a5,DT_in:=#DT_in,TS:=#tx);
         #x5 := #s5;
         #cnt := #cnt + 1;
         #ESR_Flag := TRUE;
     END_IF;
     IF #cnt < 4 AND #s6 <> #x6 AND ((BYTE_TO_INT(#s6) < 100) OR (BYTE_TO_INT(#s6) > 99 AND BYTE_TO_INT(#s6) < 200 AND BYTE_TO_INT(#Mode) >= 2) OR (BYTE_TO_INT(#s6) > 199 AND #Mode = 3)) THEN
         #ESR_Out[#cnt] := "STATUS_TO_ESR"(status:=#s6,adress:=#a6,DT_in:=#DT_in,TS:=#tx);
         #x6 := #s6;
         #cnt := #cnt + 1;
         #ESR_Flag := TRUE;
     END_IF;
     IF #cnt < 4 AND #s7 <> #x7 AND ((BYTE_TO_INT(#s7) < 100) OR (BYTE_TO_INT(#s7) > 99 AND BYTE_TO_INT(#s7) < 200 AND BYTE_TO_INT(#Mode) >= 2) OR (BYTE_TO_INT(#s7) > 199 AND #Mode = 3)) THEN
         #ESR_Out[#cnt] := "STATUS_TO_ESR"(status:=#s7,adress:=#a7,DT_in:=#DT_in,TS:=#tx);
         #x7 := #s7;
         #cnt := #cnt + 1;
         #ESR_Flag := TRUE;
     END_IF;


   (* revision history
   hm  26. jan 2007    rev 1.0
     original version

   hm  17. sep 2007  rev 1.1
     replaced time() with T_PLC_MS() for compatibility reasons

   hm  1. dec. 2009  rev 1.2
     changed esr_out to be I/O


   *)
END_FUNCTION_BLOCK

FUNCTION_BLOCK "STIME"   // FB64, SCL
TITLE = STIME
{ S7_Optimized_Access := 'FALSE' }
AUTHOR : dalbi
FAMILY : MEASURE
NAME : STIME
VERSION : 1.4
// this function block makes sure that the timer of a siemens sps counts from 0 - 2^32-1.
   VAR_OUTPUT
      tx : DWord;
      at_tx AT tx : Array[0..31] of Bool;
   END_VAR
   VAR
      last_time : DWord;
      bit31 : Bool;
      init : Bool := TRUE;
   END_VAR
   VAR_TEMP
      TOP_SI : Struct
         EV_CLASS : Byte;
         EV_NUM : Byte;
         PRIORITY : Byte;
         NUM : Byte;
         TYP2_3 : Byte;
         TYP1 : Byte;
         ZI1 : Word;
         ZI2_3 : DWord;
      END_STRUCT;
      START_UP_SI : Struct
         EV_CLASS : Byte;
         EV_NUM : Byte;
         PRIORITY : Byte;
         NUM : Byte;
         TYP2_3 : Byte;
         TYP1 : Byte;
         ZI1 : Word;
         ZI2_3 : DWord;
      END_STRUCT;
      ERR : Int;
   END_VAR
BEGIN


   (* this FB is only necessary for siemens sps
   the siemens sps timer counts from 0 to 2^31-1 and starts at 0 sfter overrun.
   this means that the bit 31 (the highest bit ) will never be used and therefore
   a problem arises when t2 - t1 is checked.
   t2 - t1 is always valid also in an timer overrun situation where the time t1 is very high and t2 is very low.
   the result of the subtraction t2 - t1 however is still valid.
   this calculation does not work for soiemens because the highest bit is not used.

   this module stores the highest bit, changes the highest bit at every overrun occurence and stuffs ther highest bit in the output.
   the output is then used by t_plc_us and t_plc_ms.

   the correction needs and fb and not a function because the value of the highest bit has to be stored.

   do never use this function block in a codesys environment. the timer in codesys is correct and runs from 0 to 2^32-1
   *)

   (* read actual startup info *)
   (* OB1_SCAN_1  BYTE  -  B#16#01: Abschluss des Neustarts (Warmstarts)
                        -  B#16#02: Abschluss des Wiederanlaufs
                        -  B#16#03: Abschluss des freien Zyklus
                        -  B#16#04: Abschluss des Kaltstarts
                        -  B#16#05: Erster OB 1-Zyklus der neuen Master-CPU nach 
                                    Master-Reserve-Umschaltung und STOP des 
                                    bisherigen Masters *)

   #ERR := RD_SINFO (TOP_SI => #TOP_SI, START_UP_SI => #START_UP_SI);

   (* reset last_time on system startup *)
   IF #TOP_SI.EV_NUM = 1 OR #TOP_SI.EV_NUM = 2 OR #TOP_SI.EV_NUM = 4 OR NOT #init THEN 
       #last_time := 0;
       #bit31 := false;
       #init := true;
   END_IF;

   (* read the system timer *)
   #tx := DINT_TO_DWORD(T_CONV(TIME_TCK()));

   (* check for overrun *)
   IF DWORD_TO_DINT(#tx) < DWORD_TO_DINT(#last_time) THEN
       (* an overrun has occured, change the value of the highest bit *)
       #bit31 := NOT #bit31;
   END_IF;

   (* stuff the highest bit into the timer value *)
   #at_tx[7] := #bit31;

   (* remember the last system time for the next overrun check *)
   #last_time := #tx;


   (* revision history
   DA  14.9.2007 rev 1.0
     original version

   DA  24.2.2008 rev 1.1
     added self reset on system startup

   DA   2.5.2008 rev 1.2
     corect a problem running under OB35

   DA  12.3.2009 rev 1.3
     corect a problem run on different CPUs

   DA  22.12.2009 rev 1.4
     corect a problem on startup
   *)
END_FUNCTION_BLOCK

FUNCTION "OSCAT_VERSION" : DWord   // FC50, SCL
TITLE = OSCAT_VERSION
{ S7_Optimized_Access := 'FALSE' }
AUTHOR : hugo
FAMILY : OTHER
NAME : OSCAT
VERSION : 1.1
// oscat_version returns the version number in dword format
// 132 is library version 1.32
// if IN = true then the release date will be returned
   VAR_INPUT
      in : Bool;
   END_VAR
BEGIN


   IF #in THEN
       #OSCAT_VERSION := DINT_TO_DWORD(T_CONV(D#2011-05-04));
   ELSE
       #OSCAT_VERSION := DW#16#0000_0332;
   END_IF;


   (* revision history
   hm  6. oct 2006 rev 1.0
     original version

   hm  16. dec 2007  rev 1.1
     added possibility to return date and version depoending on in.

   *)
END_FUNCTION

FUNCTION "STATUS_TO_ESR" : "ESR_DATA"   // FC51, SCL
TITLE = STATUS_TO_ESR
{ S7_Optimized_Access := 'FALSE' }
AUTHOR : hugo
FAMILY : OTHER
NAME : STAT_ESR
VERSION : 1.0
// status_to_esr creates esr data from a status byte.
// 
// uses: ESR_DATA [UDT8]
   VAR_INPUT
      status : Byte;
      adress : String[254];
      DT_in : Date_And_Time;
      TS : Time;
   END_VAR
   VAR_TEMP
      tstatus_to_ESR : "ESR_DATA";
   END_VAR
BEGIN


     IF BYTE_TO_INT(#status) < 100 THEN
         #tstatus_to_ESR.TYP := 1;
     ELSIF BYTE_TO_INT(#status) < 200 THEN
         #tstatus_to_ESR.TYP := 2;
     ELSE
         #tstatus_to_ESR.TYP := 3;
     END_IF;
     #tstatus_to_ESR.ADRESS:= #adress;
     #tstatus_to_ESR.DS := #DT_in;
     #tstatus_to_ESR.TS := #TS;
     #tstatus_to_ESR.DATA[0] := #status;

     #STATUS_TO_ESR := #tstatus_to_ESR;
END_FUNCTION

FUNCTION "INC1" : Int   // FC53, SCL
TITLE = INC1
{ S7_Optimized_Access := 'FALSE' }
AUTHOR : hugo
FAMILY : MATH
NAME : INC1
VERSION : 1.2
// This is a increment function which increments the variable X by 1 and if M is reached, it begins with 0 again.
// _inc1(3,X) will generate 0,1,2,3,0,1,.....
   VAR_INPUT
      X : Int;
      N : Int;
   END_VAR
BEGIN


   IF #X >= #N - 1 THEN
       #INC1 := 0;
   ELSE
       #INC1 := #X + 1;
   END_IF;


   (* this elegant version is 50% slower
   INC1 := X := (x + 1) MOD N;
   *)



   (* revision history
   hm  13. oct. 2008   rev 1.0
       original version

   hm  22. oct. 2008   rev 1.1
       added statement to return value for compatibility reasons

   hm  23. feb. 2009   rev 1.2
       when inc1 is called with X >= N inc will continue with 0
   *)
END_FUNCTION

FUNCTION "T_PLC_MS" : DWord   // FC64, SCL
TITLE = T_PLC_MS
{ S7_Optimized_Access := 'FALSE' }
AUTHOR : hugo
FAMILY : MEASURE
NAME : T_PLC_MS
VERSION : 1.2
// T_PLC_MS reads the internal PLC timer and return the time, it has the advantage to be able to set a debug mode 
// and speed up the counter to test the plc timer overrun which occurs every 50 days respectively 25 days at siemens S7
// this routine also allows to correct the behavior of s7 where the internal plc counter will not count all 32 bits.
// 
// uses: STIME [FB64],IDB_STIME [DB64]
BEGIN


   "IDB_STIME"(); 
   #T_PLC_MS := "IDB_STIME".tx; 
   (* hier muss die korrektur für step7 stattfinden
   plctime muss den vollen wertebereich von time ausnutzen:
   wenn bei step7 time -24tage bis plus 24 tage ist dann muss der timer auch beim überlauf auf -24tage springen 
   und auf keinen fall auf 0 !!!!
   für siemens muss ein weiterer fb im main eingebunden werden der sicherstellt das alle 32 bits durchgezählt werden.
   es kann nur ein fb sein den er muss sich das oberste (32te) bit merken.
   oder etwa spring s7 bei überlauf auf -24 tage????? dann wäre keine korrektur nötig.
   *)
   IF "debug" THEN
       #T_PLC_MS := DINT_TO_DWORD((DWORD_TO_DINT(SHL(IN:=#T_PLC_MS,N:="N") OR SHL(IN:=DWORD#1,N:="N"))-1) + DWORD_TO_DINT("offset_1"));
   END_IF;


   (* revision history
   hm  14.9.2007   rev 1.0
       original version

   hm  12. nov 2007    rev 1.1
       added temporaray variable tx because some compilers could not handle time() as an argument

   hm  16. nov. 2008   rev 1.2
       initialized constants with 0 for compatibility reasons
   *)
END_FUNCTION

FUNCTION "DIFFER" : Bool   // FC73, SCL
TITLE = DIFFER
{ S7_Optimized_Access := 'FALSE' }
AUTHOR : hugo
FAMILY : MATH
NAME : DIFFER
VERSION : 1.1
// this function checks if in1 differs more then x from in2
// the output is true if in1 < in2 - x or in1 > in2 + X
   VAR_INPUT
      in1 : Real;
      in2 : Real;
      X : Real;
   END_VAR
BEGIN


   #DIFFER := ABS(#in1 - #in2) > #X;

   (* revision history
   hm    8. oct 2006   rev 1.0
     original version

   hm    16. mar 2008  rev 1.1
     improverd code for performance

   *)
END_FUNCTION

// ===== PLC "String"  Unspecific CPU S7 300 =====

VAR_GLOBAL CONSTANT   // PLC tag table "STEP7 classic symbols"
   "MTH_OFS1" : Int := 0;
   "MTH_OFS2" : Int := 31;
   "MTH_OFS3" : Int := 59;
   "MTH_OFS4" : Int := 90;
   "MTH_OFS5" : Int := 120;
   "MTH_OFS6" : Int := 151;
   "MTH_OFS7" : Int := 181;
   "MTH_OFS8" : Int := 212;
   "MTH_OFS9" : Int := 243;
   "MTH_OFS10" : Int := 273;
   "MTH_OFS11" : Int := 304;
   "MTH_OFS12" : Int := 334;
   "FILL_FC235" : Char := '0';   // MigChange: FILL
   "BLANK" : Char := ' ';
END_VAR

DATA_BLOCK "SETUP"   // DB1
TITLE = SETUP
{ S7_Optimized_Access := 'FALSE' }
AUTHOR : oscat
FAMILY : CONSTANT
NAME : DBSETUP
VERSION : 1.0
   VAR
      EXTENDED_ASCII : Bool := TRUE;
      CHARNAMES : Array[1..4] of String[253];
      MTH_OFS : Array[1..12] of Int;
      DECADES : Array[0..8] of Real;
   END_VAR
BEGIN
   CHARNAMES[1] := ';"&quot;&&amp;<&lt;>&gt;€&euro; &nbsp;¡&iexcl;¢&cent;£&pound;¤&curren;¥&yen;¦&brvbar;§&sect;¨&uml;©&copy;ª&ordf;«&laquo;¬&not;­&shy;®&reg;¯&macr;°&deg;±&plusmn;²&sup2;³&sup3;´&acute;µ&micro;¶&para;·&middot;¸&cedil;¹&sup1;º&ordm;»&raquo;¼&frac14;Û&Ucirc;';
   CHARNAMES[2] := ';¾&frac34;¿&iquest;À&Agrave;Á&Aacute;Â&Acirc;Ã&Atilde;Ä&Auml;Å&Aring;Æ&AElig;Ç&Ccedil;È&Egrave;É&Eacute;Ê&Ecirc;Ë&Euml;Ì&Igrave;Í&Iacute;Î&Icirc;Ï&Iuml;Ð&ETH;Ñ&Ntilde;Ò&Ograve;Ó&Oacute;Ô&Ocirc;Õ&Otilde;Ö&Ouml;×&times;Ø&Oslash;Ù&Ugrave;Ú&Uacute;½&frac12;';
   CHARNAMES[3] := ';Ü&Uuml;Ý&Yacute;Þ&THORN;ß&szlig;à&agrave;á&aacute;â&acirc;ã&atilde;ä&auml;å&aring;æ&aelig;ç&ccedil;è&egrave;é&eacute;ê&ecirc;ë&euml;ì&igrave;í&iacute;î&icirc;ï&iuml;ð&eth;ñ&ntilde;ò&ograve;ó&oacute;ô&ocirc;õ&otilde;ö&ouml;÷&divide;ø&oslash;ù&ugrave;';
   CHARNAMES[4] := ';ú&uacute;û&ucirc;ü&uuml;ý&yacute;þ&thorn;ÿ&yuml;';
   MTH_OFS[2] := 31;
   MTH_OFS[3] := 59;
   MTH_OFS[4] := 90;
   MTH_OFS[5] := 120;
   MTH_OFS[6] := 151;
   MTH_OFS[7] := 181;
   MTH_OFS[8] := 212;
   MTH_OFS[9] := 243;
   MTH_OFS[10] := 273;
   MTH_OFS[11] := 304;
   MTH_OFS[12] := 334;
   DECADES[0] := 1.0e+0;
   DECADES[1] := 1.0e+1;
   DECADES[2] := 1.0e+2;
   DECADES[3] := 1.0e+3;
   DECADES[4] := 1.0e+4;
   DECADES[5] := 1.0e+4;
   DECADES[6] := 1.0e+5;
   DECADES[7] := 1.0e+6;
   DECADES[8] := 1.0e+7;
END_DATA_BLOCK

